// TIA Portal project "Parsing_migrated" (V16)

(* hardware
DEVICE "S71500/ET200MP station_1"  S7-1500 station
   slot 0: "Rail_0"  Rack  6ES7 590-1***0-0AA0
   slot 1: "PLC_1"  CPU 1515TF-2 PN  6ES7 515-2UM01-0AB0  V2.8
      slot 3: "CPU display_1"  6ES7591-1BA00-0AA0
      slot 32768: "PROFINET interface_1"  X1
         slot 32769: "Port_1"  X1 P1
         slot 32770: "Port_2"  X1 P2
      slot 33024: "PROFINET interface_2"  X2
         slot 33025: "Port_1"  X2 P1
      slot 34817: "Virtual CP interface port_1"  Virtual CP interface port  Virtual CP interface port
DEVICE "HMI_1"  KTP700F Mobile
   slot 0: "HMI_1"  KTP700F Mobile  6AV2 125-2GB23-0AX0  16.0.0.0
   slot 1: "HMI_RT_1"  KTP700F Mobile  6AV2 125-2GB23-0AX0  16.0.0.0
   slot 5: "HMI_1.IE_CP_1"  PROFINET Interface  16.0.0.0
      slot 1: "PROFINET Interface_1"  PROFINET Interface
         slot 1: "Port_1"  Port
DEVICE "SINAMICS S_1"  AcxSinamics.Device.2x.S210
   slot 0: "Left"  S210 PN  6SL3210-5HB10-1xFx  V5.2
      slot 1: "PROFINET interface"  PROFINET
      slot 3: " Ethernet commissioning interface"  LAN
   slot 0: "Drive control"  S210 PN
      slot 200: "Motor_Module_2"  Drive control  6SL3210-5HB10-1xFx
      slot 300: "SMIXX_3"  Drive control  1FK2102-1AG0x-xDAx
      slot 400: "Encoder_4"  Drive control  1FK2102-1AG0x-xDAx
      slot 1000: "Motor_SMI_5"  Drive control  1FK2102-1AG0x-xDAx
DEVICE "SINAMICS S_2"  AcxSinamics.Device.2x.S210
   slot 0: "Right"  S210 PN  6SL3210-5HB10-1xFx  V5.2
      slot 1: "PROFINET interface"  PROFINET
      slot 3: " Ethernet commissioning interface"  LAN
   slot 0: "Drive control"  S210 PN
      slot 200: "Motor_Module_2"  Drive control  6SL3210-5HB10-1xFx
      slot 300: "SMIXX_3"  Drive control  1FK2102-1AG0x-xDAx
      slot 400: "Encoder_4"  Drive control  1FK2102-1AG0x-xDAx
      slot 1000: "Motor_SMI_5"  Drive control  1FK2102-1AG0x-xDAx
*)

// ===== PLC "PLC_1"  CPU 1515TF-2 PN =====

VAR_GLOBAL   // PLC tag table "Default tag table"
   "PositioningAxis_Left_Actor_Interface_AddressIn" AT %I276.0 : "PD_TEL105_IN";
   "PositioningAxis_Left_Actor_Interface_AddressOut" AT %Q276.0 : "PD_TEL105_OUT";
   "PositioningAxis_Right_Actor_Interface_AddressIn" AT %I256.0 : "PD_TEL105_IN";
   "PositioningAxis_Right_Actor_Interface_AddressOut" AT %Q256.0 : "PD_TEL105_OUT";
   "actuator" AT %Q0.0 : Bool;
END_VAR

VAR_GLOBAL CONSTANT   // PLC tag table "LKinCtrl_PLC_Tags"
   "LKINCTRL_MC_MOVELINEARABS" : Int := 1;   // cmdType for linear absolute command
   "LKINCTRL_MC_MOVELINEARREL" : Int := 2;   // cmdType for linear relative command
   "LKINCTRL_MC_MOVECIRCULARABS" : Int := 3;   // cmdType for circular absolute command
   "LKINCTRL_MC_MOVECIRCULARREL" : Int := 4;   // cmdType for circular relative command
   "LKINCTRL_NO_OF_PATHDATA_PREBUFFER_ELEMENTS" : Int := 5;   // number of PreBuffer elements
   "LKINCTRL_NO_OF_START_EXECUTE_CMDS" : Int := 5;   // number of cmds to be buffered in first cycle
   "LKINCTRL_NO_OF_SEQ_EXECUTE_CMDS" : Int := 1;   // number of cmds to be buffered after first cycle
   "LKINCTRL_PI" : LReal := 3.1415926535897932846264;   // constant value for pi
   "LKINCTRL_NO_OF_CMD_SETFLAGS" : Int := 3;   // number of Boolean flags per command
   "LKINCTRL_LENGTH_OF_CMDPOINT_NAME" : Int := 10;   // length of point name
   "LKINCTRL_FM_SET_BEFORE_AND_NO_RESET" : USInt := 1;   // set flag before cmd and no reset
   "LKINCTRL_FM_SET_BEFORE_AND_RESET_AFTER" : USInt := 2;   // set flag before cmd and reset after
   "LKINCTRL_FM_SET_BEFORE_AND_RESET_AFTER_ONE_CYCLE" : USInt := 3;   // set flag before cmd and reset after one cycle
   "LKINCTRL_FM_SET_BEFORE_AND_NO_RESET_AND_WAIT_FOR_ACKNOWLEDGE" : USInt := 5;   // set flag before cmd and wait for external reset
   "LKINCTRL_FM_SET_AFTER_AND_NO_RESET" : USInt := 11;   // set flag after cmd and no reset
   "LKINCTRL_FM_SET_AFTER_AND_RESET_AFTER_ONE_CYCLE" : USInt := 13;   // set flag after cmd and reset after one cycle
   "LKINCTRL_FM_SET_AFTER_AND_NO_RESET_AND_WAIT_FOR_ACKNOWLEDGE" : USInt := 15;   // set flag after cmd and wait for external reset
   "LKINCTRL_FM_SET_AT_REMAINING_DISTANCE" : USInt := 10;   // set flag at remaining distance
   "LKINCTRL_FM_DISTANCE_TOLERANCE" : LReal := 0.01;   // tolerance for flagmode 10
   "LKINCTRL_NO_OF_SETFLAGS_BUFFER_ELEMENTS" : Int := 15;   // set as double of LKINCTRL_NO_OF_PATHDATA_PREBUFFER_ELEMENTS
   "LKINCTRL_COMP_LEFT" : Int := 1;   // tool radius compensation to the left
   "LKINCTRL_COMP_RIGHT" : Int := 2;   // tool radius compensation to the right
   "LKINCTRL_OUTER_CORNER" : Int := 1;   // Outer corner (linear / linear intersection)
   "LKINCTRL_INNER_CORNER" : Int := 2;   // Inner corner (linear / linear intersection)
   "LKINCTRL_CONFIG_END_OFFSET_COMP" : Int := 40;   // cmdType for ending offset compensation
   "LKINCTRL_CONFIG_START_OFFSET_COMP_LEFT" : Int := 41;   // cmdType for starting offset compensation left
   "LKINCTRL_NO_OF_PATHDATA_ELEMENTS" : Int := 20;   // length of LKinCtrl_typePathData
   "LKINCTRL_CMD_WAIT_TIME" : Int := 100;   // cmdType for wait time command
   "LKINCTRL_CONFIG_START_OFFSET_COMP_RIGHT" : Int := 42;   // cmdType for starting offset compensation right
   "LKINCTRL_LENGTH_OF_OFFSET_NAME" : Int := 10;   // length of offset name
   "LKINCTRL_NO_OF_OFFSETS" : Int := 3;   // number of configurable offsets
   "LKINCTRL_PATHDATA_TYPE_REDUCED" : USInt := 1;   // constant for PathData type "reduced"
   "LKINCTRL_PATHDATA_TYPE_NORMAL" : USInt := 2;   // constant for PathData type "normal"
   "LKINCTRL_PATHDATA_TYPE_ADVANCED" : USInt := 3;   // constant for PathData type "advanced"
   "LKINCTRL_NO_OF_PATHDATA_ELEMENTS_ADVANCED" : Int := 20;   // length of LKinCtrl_typePathData_advanced
   "LKINCTRL_NO_OF_PATHDATA_ELEMENTS_REDUCED" : Int := 10;   // length of LKinCtrl_typePathData_reduced
   "LKINCTRL_NO_OF_VALID_BITS" : Int := 4;   // number of valid bits in PathDataElement_advanced
   "LKINCTRL_CIRCMODE_GCODE" : Int := 3;   // circMode used in GCode
   "LKINCTRL_CMD_FLAG_ONLY" : Int := 0;   // cmdType for flagOnly command (no motion)
   "LKINCTRL_FM_DEACTIVATED" : USInt := 0;   // flag deactiavted
   "LKINCTRL_NO_OF_CMD_VALUEFLAGS" : Int := 3;   // number of LREAL flags per command
   "LKINCTRL_NO_OF_LAST_SETFLAG" : Int := 5;   // number of set flags at MovePath FB
   "LKINCTRL_NO_OF_LAST_VALUEFLAG" : Int := 5;   // number of value flags at MovePath FB
   "LKINCTRL_LENGTH_OF_PATHDATA_NAME" : Int := 15;   // length of PathData name
   "LKINCTRL_MC_MOVEDIRECTABS" : Int := 5;   // cmdType for move direct absolute command
   "LKINCTRL_MC_MOVEDIRECTREL" : Int := 6;   // cmdType for move direct relative command
   "LKINCTRL_NO_OF_CONVEYOR" : Int := 3;   // number of configurable offsets
   "LKINCTRL_MC_TRACKCONVEYORBELT" : Int := 10;   // cmdType for track conveyor belt command
END_VAR

VAR_GLOBAL CONSTANT   // PLC tag table "MC_Constants"
   "BM_BUFFERED" : Int := 1;   // Buffer mode 1: Standstill between motions
   "BM_BLENDING_LOW" : Int := 2;   // Buffer mode 2: Blending with lower velocity
   "BM_BLENDING_HIGH" : Int := 5;   // Buffer mode 5: Blending with higher velocity
   "DA_DEFAULT" : Int := -1;   // Dynamic adaption -1: Use default
   "DA_DEACTIVATED" : Int := 0;   // Dynamic adaption 0: Deactivated
   "DA_WITH_VARIABLE_LIMITS" : Int := 1;   // Dynamic adaption 1: With segmentation of path
   "DA_WITH_CONSTANT_LIMITS" : Int := 2;   // Dynamic adaption 2: No segmentation of path
   "SM_ACTIVE_DYNAMICS" : Int := 0;   // Stop mode 0: Stop with active dynamics
   "SM_MAX_DYNAMICS" : Int := 1;   // Stop mode 1: Stop with maximum dynamics
   "PC_POSITIVE" : Int := 0;   // Path choice 0: Shorter positive circle segment
   "PC_LONG_RUN_POSITIVE" : Int := 2;   // Path choice 2: Longer positive circle segment
   "PC_LONG_RUN_NEGATIVE" : Int := 3;   // Path choice 3: Longer negative circle segment
   "CP_XZ" : Int := 0;   // Circle plane 0: Circle in X-Z plane
   "CP_YZ" : Int := 1;   // Circle plane 1: Circle in Y-Z plane
   "CP_XY" : Int := 2;   // Circle plane 2: Circle in X-Y plane
   "CM_BORDER" : Int := 0;   // Circle mode 0: "EndPoint" + "AuxPoint" parameter defines a point on circular path
   "CM_CENTER" : Int := 1;   // Circle mode 1: "Arc" + "AuxPoint" defines circle center
   "CM_RADIUS" : Int := 2;   // Circle mode 2: "Radius" + "EndPoint" parameters define the circle segment
   "IM_ACTIVE_DYNAMICS" : Int := 0;   // Interrupt mode 0: Interrupt with active dynamics
   "IM_MAX_DYNAMICS" : Int := 1;   // Interrupt mode 1: Interrupt with maximum dynamics
   "DIRA_POSITIVE" : Int := 1;   // Orientation direction 1: Positive direction
   "DIRA_NEGATIVE" : Int := 2;   // Orientation direction 2: Negative direction
   "DIRA_SHORTEST" : Int := 3;   // Orientation direction 3: Shortest direction
   "CS_WCS" : Int := 0;   // Coordinate system 0: World coordinate system (WCS)
   "CS_OCS1" : Int := 1;   // Coordinate system 1: Object coordinate system 1 (OCS[1])
   "CS_OCS2" : Int := 2;   // Coordinate system 2: Object coordinate system 2 (OCS[2])
   "CS_OCS3" : Int := 3;   // Coordinate system 3: Object coordinate system 3 (OCS[3])
   "PC_NEGATIVE" : Int := 1;   // Path choice 1: Shorter negative circle segment
   "CS_MCS" : Int := 100;   // Coordinate system 100: Machine coordinate system (axis values)
   "LC_DEFAULT" : DWord := 16#FFFFFFFF;   // LinkConstellation: Default to keep link constellation of kinematics
   "PM_ABS_ABS" : DInt := 1;   // PositionMode 1: Interpretation of cartesian orientation as absolute (only effective for absolute MoveDirect commands)
   "PM_ABS_REL" : DInt := 2;   // PositionMode 2: Interpretation of cartesian orientation as relative (only effective for absolute MoveDirect commands)
END_VAR

VAR_GLOBAL CONSTANT   // PLC tag table "LKinLang_Configuration"
   "LKINLANG_FIRST_INDEX_LINE_BUFFER" : Int := 1;   // First index of the line buffer
   "LKINLANG_LAST_INDEX_LINE_BUFFER" : Int := 20;   // Last index of the line buffer
   "LKINLANG_LENGTH_OF_ASCII_LINE_STRING" : UDInt := 128;   // Maximum number of ASCII characters in one line (without CR/LF)
   "LKINLANG_LENGTH_OF_TOKEN_STRING" : Int := 20;   // Maximum string length of one token
   "LKINLANG_MAX_NUMBER_OF_TOKEN_PER_LINE" : Int := 50;   // Maximum number of token per line
   "LKINLANG_MAX_NUMBER_OF_PARAMETERS_PER_LINE" : Int := 25;   // Maximum number of parameters in one line
   "LKINLANG_MAX_NUMBER_OF_PARAMETERS" : Int := 125;   // Maximum number of configured language parameters (G1,G2,...)
   "LKINLANG_NUMBER_OF_SEPARATORS" : Int := 15;   // Maximum number of separators
   "LKINLANG_NUMBER_OF_MERGERS" : Int := 10;   // Maximum number of mergers
   "LKINLANG_NUMBER_OF_FOLLOW_VALUES" : Int := 4;   // Maximum number of follow values for one command
   "LKINLANG_NUMBER_OF_CONDITIONS" : Int := 50;   // Maximum number of conditions for one command
   "LKINLANG_NUMBER_OF_REPLACEMENTS" : Int := 10;   // Maximum number of replacements
   "LKINLANG_NUMBER_OF_LABELS" : Int := 20;   // Maximum number of labels
   "LKINLANG_NUMBER_OF_STACK_ELEMENTS" : Int := 20;   // Maximum number of stack elements
   "LKINLANG_NUMBER_OF_HIERARCHICLEVEL" : Int := 60;   // Maximum number of hierarchic level changes
   "LKINLANG_NUMBER_OF_SUBPROGRAMS" : Int := 10;   // Maximum number of subprograms
   "LKINLANG_NUMBER_OF_VAR_REFS" : Int := 20;   // Maximum number of variable references
   "LKINLANG_NUMBER_OF_INTERFACE_BOOL" : Int := 5;   // Maximum number of boolean interface variables
   "LKINLANG_NUMBER_OF_INTERFACE_DINT" : Int := 10;   // Maximum number of DInt interface variables
   "LKINLANG_NUMBER_OF_INTERFACE_LREAL" : Int := 20;   // Maximum number of LReal interface variables
   "LKINLANG_NUMBER_OF_LOCAL_BOOL" : Int := 10;   // Maximum number of boolean local variables
   "LKINLANG_NUMBER_OF_LOCAL_DINT" : Int := 10;   // Maximum number of DInt local variables
   "LKINLANG_NUMBER_OF_LOCAL_LREAL" : Int := 10;   // Maximum number of LReal local variables
   "LKINLANG_LANGPACK_GCODE" : Int := 1;   // Select GCode language package
   "LKINLANG_LANGPACK_USER" : Int := 2;   // Select user defined language package
END_VAR

VAR_GLOBAL CONSTANT   // PLC tag table "LKinLang_Constants"
   "LKINLANG_PRIO_UNRELEVANT" : Int := 0;   // Lowest parameter priority
   "LKINLANG_PRIO_DEFAULT" : Int := 1;   // Normal parameter priority
   "LKINLANG_PRIO_DEFINED" : Int := 2;   // High parameter priority
   "LKINLANG_PRIO_CONSTANT" : Int := 3;   // Highest parameter priority
   "LKINLANG_MOTION_CMD" : DWord := 2#0000_0001;   // Parameter property: Motion command
   "LKINLANG_ABSOLUTE_POSITION" : DWord := 2#0010_0000;   // Parameter property: Switch to absolute positioning
   "LKINLANG_RELATIVE_POSITION" : DWord := 2#0100_0000;   // Parameter property: Switch to relative positioning
   "LKINLANG_CMD_MODAL" : DWord := 2#0000_0010;   // Parameter property: Modal until change of motion command
   "LKINLANG_PRG_MODAL" : DWord := 2#0000_0100;   // Parameter property: Modal for complete program
   "LKINLANG_CHECK_LIMITS" : DWord := 2#0000_1000;   // Parameter property: Check limits for parameter
   "LKINLANG_EQUATION" : DWord := 2#0001_0000;   // Parameter property: Math expressions allowed
   "LKINLANG_CONDITION_IN_LINE" : DInt := 1;   // Condition check: Condition must be set in same line
   "LKINLANG_CONDITION_IN_COMMAND" : DInt := 2;   // Condition check: Condition must be set in same motion command
   "LKINLANG_CONDITION_IN_PROGRAM" : DInt := 3;   // Condition check: Condition must be set in program before
   "LKINLANG_FILE_STATE_RUNNING" : DInt := 200;   // File status: Program in execution
   "LKINLANG_FILE_STATE_STOPPED" : DInt := 90;   // File status: Program stopped
   "LKINLANG_FILE_STATE_EDITING" : DInt := 20;   // File status: Program is edited
   "LKINLANG_FILE_STATE_LOADING" : DInt := 10;   // File status: Program is being loaded from MMC
   "LKINLANG_FILE_STATE_RUNNING_LOADING" : DInt := 300;   // File status: Program is executed and loaded simultaneously
   "LKINLANG_FILE_STATE_SAVING" : DInt := 30;   // File status: Program is being saved
   "LKINLANG_FILE_STATE_IDLE" : DInt := 100;   // File status: Program is ready
   "LKINLANG_FILE_STATE_SAVE_REQUESTED" : DInt := 40;   // File status: Program saving is requested
   "LKINLANG_VAR_TYPE_LOCAL_BOOL" : Int := 1;   // Type constant for local boolean variables
   "LKINLANG_VAR_TYPE_LOCAL_DINT" : Int := 2;   // Type constant for local integer variables
   "LKINLANG_VAR_TYPE_LOCAL_LREAL" : Int := 3;   // Type constant for local real variables
   "LKINLANG_VAR_TYPE_INTERFACE_BOOL" : Int := 101;   // Type constant for boolean interface variables
   "LKINLANG_VAR_TYPE_INTERFACE_DINT" : Int := 102;   // Type constant for integer interface variables
   "LKINLANG_VAR_TYPE_INTERFACE_LREAL" : Int := 103;   // Type constant for real interface variables
   "LKINLANG_SYNTAX_CHECK_OFF" : USInt := 0;   // Constant for syntax check: No check before writing commands
   "LKINLANG_SYNTAX_CHECK_ONLY" : USInt := 1;   // Constant for syntax check: Only check; no writing of commands
   "LKINLANG_SYNTAX_CHECK_AND_EXECUTE" : USInt := 2;   // Constant for syntax check: Check before and write commands after check
   "LKINLANG_ENTRY_TYPE_IF" : Int := 10;   // Stack entry type IF
   "LKINLANG_ENTRY_TYPE_ELSE" : Int := 11;   // Stack entry type ELSE
   "LKINLANG_ENTRY_TYPE_ENDIF" : Int := 12;   // Stack entry type ENDIF
   "LKINLANG_ENTRY_TYPE_WHILE" : Int := 20;   // Stack entry type WHILE
   "LKINLANG_ENTRY_TYPE_ENDWHILE" : Int := 22;   // Stack entry type ENDWHILE
   "LKINLANG_ENTRY_TYPE_FOR" : Int := 30;   // Stack entry type FOR
   "LKINLANG_ENTRY_TYPE_ENDFOR" : Int := 32;   // Stack entry type ENDFOR
   "LKINLANG_ENTRY_TYPE_SUB" : Int := 40;   // Stack entry type SUB
END_VAR

// folder: LKinCtrl_Types

TYPE "LKinCtrl_typeFrame"
   STRUCT
      x : LReal;   // Translation in x
      y : LReal;   // Translation in y
      z : LReal;   // Translation in z
      "a" : LReal;   // Rotation around z axis
      "b" : LReal;   // Rotation around y axis
      c : LReal;   // Roataion around x axis
   END_STRUCT;
END_TYPE

TYPE "LKinCtrl_typePathDataElement_advanced"
VERSION : 0.1
   STRUCT
      cmdType : Int := -1;   // 1: MoveLinAbs; 2: MoveLinRel; 3: MoveCircAbs; 4: MoveCircRel; 5: MoveDirectAbs; 6: MoveDirectRel; 10: TrackConveyorBelt; 100: WaitTime; 40/41/42: ContourOffset; 0: FlagOnlyCmd; -1: End of List
      cmdActivated : Bool := TRUE;   // (de)activation of command
      cmdName : String["LKINCTRL_LENGTH_OF_CMDPOINT_NAME"];   // name of command
      cmdCoordinates : "LKinCtrl_typePointCoordinates";   // target coordinate definition
      cmdParameters : "LKinCtrl_typePointParameter";   // additional command parameters
      setFlags : Array[1.."LKINCTRL_NO_OF_CMD_SETFLAGS"] of "LKinCtrl_typeSetFlagElement_Bool";   // flags to control actuators
      valueFlags : Array[1.."LKINCTRL_NO_OF_CMD_VALUEFLAGS"] of "LKinCtrl_typeSetFlagElement_LReal";   // value flags to control actuators
      parameterValid : Array[1..4] of Bool;   // valid bit for cartesian position parameters
   END_STRUCT;
   // parameterValid[1] := True;   // X
   // parameterValid[2] := True;   // Y
   // parameterValid[3] := True;   // Z
   // parameterValid[4] := True;   // A
   // // cmdParameters.transitionParameters : blending parameters
   // // cmdParameters.pathDynamics : dynamic settings
END_TYPE

TYPE "LKinCtrl_typeCmdLoggerElement"
VERSION : 0.1
   STRUCT
      cmdType : Int := -1;   // 1: MoveLinAbs; 2: MoveLinRel; 3: MoveCircAbs; 4: MoveCircRel; 5: MoveDirectAbs; 6: MoveDirectRel; 10: TrackConveyorBelt; 100: WaitTime; 40/41/42: ContourOffset; 0: FlagOnlyCmd; -1: End of List
      pathDataName : String["LKINCTRL_LENGTH_OF_PATHDATA_NAME"];   // name of PathData
      pathDataIdentifier : Int;   // identifier of PathData containing command
      cmdID : DInt;   // to be set to PathDataOperate[list position] by PreBuffer for identification in ExecuteBuffer
      cmdName : String[4];   // command name
      coordinateX : LReal;   // X (linear) / endPoint[1] (circular)
      coordinateY : LReal;   // Y (linear) / endPoint[2] (circular)
      coordinateZ : LReal;   // Z (linear) / endPoint[3] (circular)
      coordinateA : LReal;   // A (linear) / endPoint[4] (circular)
      coordSystem : DInt := 0;   // 0: WCS; 1: OCS[1]; 2: OCS[2]; 3: OCS[3]
      bufferMode : DInt := 1;   // 1: standstill between commands, 2: blending with lower speed; 5: blending with higher speed
      transitionParameter : LReal;   // blending distance - >0.0: configured value used; <0.0: maximum possible blending distance used
      dynVelocity : LReal;   // >0.0: configured value used; <0.0: default TO setting used
      dynAcceleration : LReal;   // >0.0: configured value used; <0.0: default TO setting used
      dynDeceleration : LReal;   // >0.0: configured value used; <0.0: default TO setting used
      dynJerk : LReal;   // >0.0: configured value used; <0.0: default TO setting used
      dynamicAdpation : DInt;   // <0.0: default TO setting used; 0: no dynamic adaption; 1: with variable limits; 2: with constant limits
      linkConstellation : DWord;   // linkConstellation (effective for MoveDirect commands only)
      positionMode : DInt;   // 1: absolute cartesian position and absolute orientation; 2: absolute cartesian position and relative orientation (effective for MoveDirect commands only)
      circMode : DInt;   // 0: auxPoint defines point on circle line; 1: auxPoint defines circle center; 2: radius and endPoint define circle segment
      auxPoint_1 : LReal;   // auxiliary point for circle definition
      auxPoint_2 : LReal;   // auxiliary point for circle definition
      auxPoint_3 : LReal;   // auxiliary point for circle definition
      pathChoice : DInt;   // circMode(0): not relevant; circMode(1): 0: pos direction; 1: neg direction; circMode(2): 0: short pos segment; 1: short neg segment; 2: long pos segment; 3: long neg segment
      circlePlane : DInt;   // circMode(0): not relevant; circMode(1+2): 0: XZ; 1: YZ; 2: XY
      radius : LReal;   // only in combination with circMode(2): radius
      arc : LReal;   // only in combination with circMode(1): arc
   END_STRUCT;
END_TYPE

TYPE "LKinCtrl_typeSetFlagElement_LReal"
VERSION : 0.1
   STRUCT
      flag : Int := -1;   // index of flag to be set
      value : LReal := 0.0;   // value for flagValue
      flagMode : USInt := 1;   // (see LKinCtrl_PLC_Tags) 0: deactivated; 1: SET_BEFORE_AND_NO_RESET; 2: SET_BEFORE_AND_RESET_AFTER; 3: SET_BEFORE_AND_RESET_AFTER_ONE_CYCLE; 5: SET_BEFORE_AND_NO_RESET_AND_WAIT_FOR_ACKNOWLEDGE; 10: LKINCTRL_FM_SET_AT_REMAINING_DISTANCE; 11: LKINCTRL_FM_SET_AFTER_AND_NO_RESET; 13: LKINCTRL_FM_SET_AFTER_AND_RESET_AFTER_ONE_CYCLE; 15: LKINCTRL_FM_SET_AFTER_AND_NO_RESET_AND_WAIT_FOR_ACKNOWLEDGE
      remainingDistance : LReal := -1.0;   // >0.0: remainingDistance
   END_STRUCT;
END_TYPE

TYPE "LKinCtrl_typeSetFlagElement_Bool"
VERSION : 0.1
   STRUCT
      flag : Int := -1;   // flag to be set
      flagMode : USInt := 1;   // (see LKinCtrl_PLC_Tags) 0: deactivated; 1: SET_BEFORE_AND_NO_RESET; 2: SET_BEFORE_AND_RESET_AFTER; 3: SET_BEFORE_AND_RESET_AFTER_ONE_CYCLE; 5: SET_BEFORE_AND_NO_RESET_AND_WAIT_FOR_ACKNOWLEDGE; 10: LKINCTRL_FM_SET_AT_REMAINING_DISTANCE; 11: LKINCTRL_FM_SET_AFTER_AND_NO_RESET; 13: LKINCTRL_FM_SET_AFTER_AND_RESET_AFTER_ONE_CYCLE; 15: LKINCTRL_FM_SET_AFTER_AND_NO_RESET_AND_WAIT_FOR_ACKNOWLEDGE
      remainingDistance : LReal := -1.0;   // >0.0: remainingDistance
   END_STRUCT;
END_TYPE

TYPE "LKinCtrl_typePointCoordinates"
VERSION : 0.1
   STRUCT
      cartesianPosition : "LKinCtrl_typeCartesianPosition";   // cartesian position
      coordSystem : DInt := 0;   // 0: WCS; 1: OCS[1]; 2: OCS[2]; 3: OCS[3] / 0: WCS; 1: OCS[1]; 2: OCS[2]; 3: OCS[3]; 100: MCS
   END_STRUCT;
END_TYPE

TYPE "LKinCtrl_typePointCoordinates_PreBuf"
VERSION : 0.1
   STRUCT
      absolutePosition : Array[1..4] of LReal;   // absolute cartesian position
      coordSystem : DInt := 0;   // 0: WCS; 1: OCS[1]; 2: OCS[2]; 3: OCS[3]
   END_STRUCT;
   // // absolutePosition[1] : X
   // // absolutePosition[2] : Y
   // // absolutePosition[3] : Z
   // // absolutePosition[4] : A
END_TYPE

TYPE "LKinCtrl_typePathDynamics"
VERSION : 0.1
   STRUCT
      velocity : LReal := -1.0;   // >0.0: configured value used; <0.0: default TO setting used; for cmdType = 100 ==> waitTime in ms
      acceleration : LReal := -1.0;   // >0.0: configured value used; <0.0: default TO setting used
      deceleration : LReal := -1.0;   // >0.0: configured value used; <0.0: default TO setting used
      jerk : LReal := -1.0;   // >0.0: configured value used; <0.0: default TO setting used
   END_STRUCT;
END_TYPE

TYPE "LKinCtrl_typePathDataElement_PreBuf"
VERSION : 0.1
   STRUCT
      cmdType : Int := -1;   // 1: MoveLinAbs; 2: MoveLinRel; 3: MoveCircAbs; 4: MoveCircRel; 5: MoveDirectAbs; 6: MoveDirectRel; 10: TrackConveyorBelt; 100: WaitTime; 40/41/42: ContourOffset; 0: FlagOnlyCmd; -1: End of List
      cmdID : DInt;   // to be set to PathDataOperate[list position] by PreBuffer for identification in ExecuteBuffer
      cmdName : String["LKINCTRL_LENGTH_OF_CMDPOINT_NAME"];   // command name
      cmdCoordinates : "LKinCtrl_typePointCoordinates_PreBuf";   // command coordinates
      cmdParameters : "LKinCtrl_typePointParameter";   // command parameters
      pathDataName : String["LKINCTRL_LENGTH_OF_PATHDATA_NAME"];   // name of PathData
      pathDataIdentifier : USInt;   // identifier of PathData
      isIntermediateCmd : Bool;   // TRUE: command is intermediate command
      setFlags : Array[1.."LKINCTRL_NO_OF_CMD_SETFLAGS"] of "LKinCtrl_typeSetFlagElement_Bool";   // flags to control actuators
      valueFlags : Array[1.."LKINCTRL_NO_OF_CMD_VALUEFLAGS"] of "LKinCtrl_typeSetFlagElement_LReal";   // value flags to control actuators
      parameterValid : Array[1..4] of Bool;   // valid bit for cartesian position parameters
   END_STRUCT;
   // parameterValid[1] := True;   // X
   // parameterValid[2] := True;   // Y
   // parameterValid[3] := True;   // Z
   // parameterValid[4] := True;   // A
END_TYPE

TYPE "LKinCtrl_typePathDescriptionElement"
   STRUCT
      pointName : String["LKINCTRL_LENGTH_OF_CMDPOINT_NAME"];   // name of point
      targetPosition : "LKinCtrl_typeCartesianPosition";   // target position
      coordSystem : DInt;   // 0: WCS; 1: OCS[1]; 2: OCS[2]; 3: OCS[3]
      blendingDistance : LReal;   // blending radius
      flags : Array[1.."LKINCTRL_NO_OF_CMD_SETFLAGS"] of "LKinCtrl_typeSetFlagElement_Bool";   // flags to control actuators
      valueFlags : Array[1.."LKINCTRL_NO_OF_CMD_VALUEFLAGS"] of "LKinCtrl_typeSetFlagElement_LReal";   // value flags to control actuators
   END_STRUCT;
END_TYPE

TYPE "LKinCtrl_typePointParameter"
VERSION : 0.1
   STRUCT
      pathDynamics : "LKinCtrl_typePathDynamics";   // dynamics settings for single command
      orientationDirection : DInt := 3;   // 1: positive direction; 2: negative direction; 3: shortest distance
      bufferMode : DInt := 1;   // 1: standstill between commands, 2: blending with lower speed; 5: blending with higher speed
      transitionParameters : Array[1..5] of LReal;   // blending distance parameters
      dynamicAdaption : DInt := -1;   // <0.0: default TO setting used; 0: no dynamic adaption; 1: with variable limits; 2: with constant limits
      moveDirectParameters : "LKinCtrl_typeMoveDirectParameter";   // parameters for MoveDirect command definition
      offsetParameters : "LKinCtrl_typeToolParameters";   // parameters for offset selection and configuration
      conveyorParameters : "LKinCtrl_typeConveyorParameter";   // parameters for conveyor selection and configuration
      circleParameters : "LKinCtrl_typeCircleParameters";   // parameters for circle command definition
   END_STRUCT;
   // transitionParameters[1] := -1.0;   // blending distance - >0.0: configured value used; <0.0: maximum possible blending distance used
   // // transitionParameters[2] : reserved, do not set
   // // transitionParameters[3] : reserved, do not set
   // // transitionParameters[4] : reserved, do not set
   // // transitionParameters[5] : reserved, do not set
END_TYPE

TYPE "LKinCtrl_typePathData_advanced"
VERSION : 0.1
   STRUCT
      pathDataName : String["LKINCTRL_LENGTH_OF_PATHDATA_NAME"];   // name of PathData
      pointers : "LKinCtrl_typeAdvPointers";   // pointers to add / retrieve cmds in PathData
      commands : Array[1.."LKINCTRL_NO_OF_PATHDATA_ELEMENTS_ADVANCED"] of "LKinCtrl_typePathDataElement_advanced";   // command list
   END_STRUCT;
END_TYPE

TYPE "LKinCtrl_typePathDataElement"
VERSION : 0.1
   STRUCT
      cmdType : Int := -1;   // 1: MoveLinAbs; 2: MoveLinRel; 3: MoveCircAbs; 4: MoveCircRel; 5: MoveDirectAbs; 6: MoveDirectRel; 10: TrackConveyorBelt; 100: WaitTime; 40/41/42: ContourOffset; 0: FlagOnlyCmd; -1: End of List
      cmdActivated : Bool := TRUE;   // (de)activation of command
      cmdName : String["LKINCTRL_LENGTH_OF_CMDPOINT_NAME"];   // name of command
      cmdCoordinates : "LKinCtrl_typePointCoordinates";   // target coordinate definition
      cmdParameters : "LKinCtrl_typePointParameter";   // additional command parameters
      setFlags : Array[1.."LKINCTRL_NO_OF_CMD_SETFLAGS"] of "LKinCtrl_typeSetFlagElement_Bool";   // flags to control actuators
      valueFlags : Array[1.."LKINCTRL_NO_OF_CMD_VALUEFLAGS"] of "LKinCtrl_typeSetFlagElement_LReal";   // value flags to control actuators
   END_STRUCT;
   // // cmdParameters.transitionParameters : blending parameters
   // // cmdParameters.pathDynamics : dynamic settings
END_TYPE

TYPE "LKinCtrl_typePathDescription"
   STRUCT
      pathDescriptionName : String[10];   // name of PathDescription
      points : Array[1.."LKINCTRL_NO_OF_PATHDATA_ELEMENTS"] of "LKinCtrl_typePathDescriptionElement";   // target points
   END_STRUCT;
END_TYPE

TYPE "LKinCtrl_typeAdvPointers"
VERSION : 0.1
   STRUCT
      addPointer : DInt := 0;   // pointer to add new comds to PathData after cmd has been executed by MovePath
      retrievePointer : DInt := 0;   // pointer to show which cmd is the next to be retrieved by MovePath
      addPointerRestarted : Bool;   // addPointer restarted after overflow
      ignoreAddPointer : Bool := true;   // addPointer not taken into account for buffering, unless set by previous data source
      bufferLocked : Bool;   // buffer locked to wait for previous data source - read data locked
      preprocessingStop : Bool;   // parser reached a preprocessing stop
   END_STRUCT;
END_TYPE

TYPE "LKinCtrl_typePointParameter_reduced"
VERSION : 0.1
   STRUCT
      pathDynamics : "LKinCtrl_typePathDynamics";   // dynamics settings for single command
      orientationDirection : DInt := 3;   // 1: positive direction; 2: negative direction; 3: shortest distance
      bufferMode : DInt := 1;   // 1: standstill between commands, 2: blending with lower speed; 5: blending with higher speed
      transitionParameters : Array[1..5] of LReal;   // blending distance parameters
      dynamicAdaption : DInt := -1;   // <0.0: default TO setting used; 0: no dynamic adaption; 1: with variable limits; 2: with constant limits
   END_STRUCT;
   // transitionParameters[1] := -1.0;   // blending distance - >0.0: configured value used; <0.0: maximum possible blending distance used
   // // transitionParameters[2] : reserved, do not set
   // // transitionParameters[3] : reserved, do not set
   // // transitionParameters[4] : reserved, do not set
   // // transitionParameters[5] : reserved, do not set
END_TYPE

TYPE "LKinCtrl_typePathData_reduced"
VERSION : 0.1
   STRUCT
      pathDataName : String["LKINCTRL_LENGTH_OF_PATHDATA_NAME"];   // name of PathData
      commands : Array[1.."LKINCTRL_NO_OF_PATHDATA_ELEMENTS_REDUCED"] of "LKinCtrl_typePathDataElement_reduced";   // command list
   END_STRUCT;
END_TYPE

TYPE "LKinCtrl_typePathData"
VERSION : 0.1
   STRUCT
      pathDataName : String["LKINCTRL_LENGTH_OF_PATHDATA_NAME"];   // name of PathData
      commands : Array[1.."LKINCTRL_NO_OF_PATHDATA_ELEMENTS"] of "LKinCtrl_typePathDataElement";   // command list
   END_STRUCT;
END_TYPE

TYPE "LKinCtrl_typePathData_PreBuf"
VERSION : 0.1
   STRUCT
      pathDataName : String["LKINCTRL_LENGTH_OF_PATHDATA_NAME"];   // name of PathData
      commands : Array[1.."LKINCTRL_NO_OF_PATHDATA_PREBUFFER_ELEMENTS"] of "LKinCtrl_typePathDataElement_PreBuf";   // command list
      addPointer : Int;   // pointer marking slot for adding of next command in PathDataPreBuffered
      retrievePointer : Int;   // pointer marking command entry to be read in PathDataPreBuffered
      addPointerRestarted : Bool;   // addPointer restarted after overflow
   END_STRUCT;
END_TYPE

TYPE "LKinCtrl_typePathDataElement_reduced"
VERSION : 0.1
   STRUCT
      cmdType : Int := -1;   // 1: MoveLinAbs; 2: MoveLinRel; 100: WaitTime; 0: FlagOnlyCmd; -1: End of List
      cmdActivated : Bool := TRUE;   // (de)activation of command
      cmdName : String["LKINCTRL_LENGTH_OF_CMDPOINT_NAME"];   // name of command
      cmdCoordinates : "LKinCtrl_typePointCoordinates";   // target coordinate definition
      cmdParameters : "LKinCtrl_typePointParameter_reduced";   // additional command parameters
      setFlags : Array[1.."LKINCTRL_NO_OF_CMD_SETFLAGS"] of "LKinCtrl_typeSetFlagElement_Bool";   // flags to control actuators
      valueFlags : Array[1.."LKINCTRL_NO_OF_CMD_VALUEFLAGS"] of "LKinCtrl_typeSetFlagElement_LReal";   // value flags to control actuators
   END_STRUCT;
END_TYPE

TYPE "LKinCtrl_typeDiagnosticsPathSelect"
TITLE = typeDiagnosticsFBTemplate
VERSION : 0.1
   STRUCT
      status : Word;   // Status of the FC or error identification when error occurred
      entryID : Int;   // identifier for false entry
   END_STRUCT;
END_TYPE

TYPE "LKinCtrl_typeExecuteKinMotionCmdDiagnostics"
VERSION : 0.1
   STRUCT
      status : Word;   // status of the FB
      faultPathDataName : String["LKINCTRL_LENGTH_OF_PATHDATA_NAME"];   // number of PathData with occurring error in PathData set
      faultSetNumber : DInt;   // number of PathData set with occurring error
      faultFBNumber : DInt;   // number of motionCommand FB with occurring error
      motionFBstatus : DWord;   // status of motion FB (internal) an error occurred in
      stateMachine : Int;   // stateMachine status
      kinematicsStatusWord : DWord;   // statusWord TO kinematics
      kinematicsErrorWord : DWord;   // errorWord TO kinematics
   END_STRUCT;
END_TYPE

TYPE "LKinCtrl_typeCircleParameters"
VERSION : 0.1
   STRUCT
      circMode : DInt := 0;   // 0: auxPoint defines point on circle line; 1: auxPoint defines circle center; 2: radius and endPoint define circle segment; 3: GCode notation (end & aux point)
      auxPoint : Array[1..3] of LReal;   // auxiliary point for circle definition
      pathChoice : DInt := 0;   // circMode(0): not relevant; circMode(1): 0: pos direction; 1: neg direction; circMode(2): 0: short pos segment; 1: short neg segment; 2: long pos segment; 3: long neg segment
      circlePlane : DInt;   // circMode(0): not relevant; circMode(1+2): 0: XZ; 1: YZ; 2: XY
      radius : LReal;   // only in combination with circMode(2): radius
      arc : LReal;   // only in combination with circMode(1): arc
   END_STRUCT;
   // // auxPoint[1] : X
   // // auxPoint[2] : Y
   // // auxPoint[3] : Z
END_TYPE

TYPE "LKinCtrl_typeMovePathDiagnostics"
VERSION : 0.1
   STRUCT
      errorID : Word;   // errorID of the FB
      pathDataName : String["LKINCTRL_LENGTH_OF_PATHDATA_NAME"];   // name of PathData an error occurred in
      cmdNumber : DInt;   // command number (in PathData) an error occurred in
      stateMovePath : DInt;   // state machine status FB
      statusSubFunction : Word;   // status of LKinCtrl_MC_ExecuteKinMotionCmd
      motionFBNumber : DInt;   // motion FB number (internal) an error occurred in
      motionFBStatus : DWord;   // status of motion FB (internal) an error occurred in
      kinematicsStatusWord : DWord;   // statusWord TO kinematics
      kinematicsErrorWord : DWord;   // errorWord TO kinematics
   END_STRUCT;
END_TYPE

TYPE "LKinCtrl_typeJogFrameDiagnostics"
VERSION : 0.1
// support: tech.team.motioncontrol@siemens.com
   STRUCT
      timeStamp : Date_And_Time;   // Time stamp at which the error occurred
      status : Word;   // Status of FB when error occurred
      stateNumber : DInt;   // State in the state machine of the FB when the error occurred
   END_STRUCT;
END_TYPE

TYPE "LKinCtrl_typeCartesianPosition"
VERSION : 0.1
   STRUCT
      x : LReal;   // X
      y : LReal;   // Y
      z : LReal;   // Z
      "a" : LReal;   // A
   END_STRUCT;
END_TYPE

TYPE "LKinCtrl_typeDynamics"
VERSION : 0.1
   STRUCT
      path : "LKinCtrl_typePathDynamics";   // Specification of the path dynamics
      orientation : "LKinCtrl_typePathDynamics";   // Specification of the orientation dynamics
      dynamicAdaption : DInt := 1;   // 0=no dynamic adaption, 1=dynamic adaptation with segmentation of the path, 2=dynamic adaptation without segmentation of the path
   END_STRUCT;
END_TYPE

TYPE "LKinCtrl_typeAuxFCDiagnostics"
TITLE = typeDiagnosticsFBTemplate
   STRUCT
      status : Word;   // Status of the FB or error identification when error occurred
      subfunctionStatus : Word;   // Status or return value of called FBs, FCs and system blocks
      axisNumber : Int;   // number of the corresponding axis the error occured in or a function effecting it
      errorDetail : UDInt;   // error detail of corresponding technology object the error occured in
      stateNumber : DInt;   // State in the state machine of the FB when the error occurred
   END_STRUCT;
END_TYPE

TYPE "LKinCtrl_typeMoveDirectParameter"
VERSION : 0.1
   STRUCT
      linkConstellation : DWord := 16#FFFFFFFF;   // linkConstellation (effective for MoveDirect commands only)
      positionMode : DInt := 1;   // 1: absolute cartesian position and absolute orientation; 2: absolute cartesian position and relative orientation (effective for MoveDirect commands only)
   END_STRUCT;
END_TYPE

TYPE "LKinCtrl_typeConfiguration"
   STRUCT
      offsetParameter : Array[1.."LKINCTRL_NO_OF_OFFSETS"] of "LKinCtrl_typeContourOffsetParameter";   // offset parameter settings
      conveyorParameter : Array[1.."LKINCTRL_NO_OF_CONVEYOR"] of "LKinCtrl_typeConveyorConfiguration";   // conveyor parameter settings
      stopMode : DInt;   // MC_GroupStop dynamics; 0: stop with dynamics of active motion job; 1: stop with maximum kinematics dynamics (dynamics adaption still effective); 10: stop with dynamics of active motion job and desync conveyor; 11: stop with maximum kinematics dynamics and desync conveyor
   END_STRUCT;
END_TYPE

TYPE "LKinCtrl_typeContourOffsetParameter"
   STRUCT
      "name" : String["LKINCTRL_LENGTH_OF_OFFSET_NAME"];   // offset name
      radius : LReal;   // offset radius
      length : LReal;   // offset length
   END_STRUCT;
END_TYPE

TYPE "LKinCtrl_typeToolParameters"
   STRUCT
      offsetParaNo : Int;   // selection of offset parameter set from configuration structure
      mainPathPlane : Int;   // main path plane for compensation
   END_STRUCT;
END_TYPE

TYPE "LKinCtrl_typeConveyorParameter"
   STRUCT
      conveyorParaNo : DInt := 1;   // selection of conveyor parameter set from configuration structure
   END_STRUCT;
END_TYPE

TYPE "LKinCtrl_typeConveyorConfiguration"
   STRUCT
      conveyorBeltAxis : DB_ANY;   // Conveyor belt axis DB
      conveyorBeltOrigin : TO_Struct_Kinematics_Frame;   // Frane to origin of conveyor belt
      initialObjectPosition : TO_Struct_Kinematics_Frame;   // Initial object position on conveyor (only x allowed)
   END_STRUCT;
END_TYPE

// folder: LKinCtrl_Types/LKinCtrl_ContOffset_Types

TYPE "LKinCtrl_typeCOff3DPoint"
VERSION : 0.1
   STRUCT
      x : LReal;   // X
      y : LReal;   // Y
      z : LReal;   // Z
   END_STRUCT;
END_TYPE

TYPE "LKinCtrl_typeCOffReturn"
   STRUCT
      returnValue : Word;   // Return value
      region : Int;   // Region type - see LKinCtrl_OffsetContour
      subBlockNumber : DInt;   // Sub function block number
      internalNumber : DInt;   // Internal number indicates the source code position
   END_STRUCT;
END_TYPE

TYPE "LKinCtrl_typeCOffPathDataIn"
   STRUCT
      currentPos : "LKinCtrl_typeCOffInCurrentPos";   // Source data - current position
      nextCommand : "LKinCtrl_typePathDataElement";   // Source data - next command
      nextButOneCommand : "LKinCtrl_typePathDataElement";   // Source data - next but one command
   END_STRUCT;
END_TYPE

TYPE "LKinCtrl_typeCOffOutNextButOneCmd"
   STRUCT
      transitionParameter : Array[1..5] of LReal;   // blending parameters
   END_STRUCT;
END_TYPE

TYPE "LKinCtrl_typeCOffCmdInInternal"
   STRUCT
      cmdType : Int := -1;   // 1: MoveLinAbs; 2: MoveLinRel; 3: MoveCircAbs; 4: MoveCircRel; 5: MoveDirectAbs; 6: MoveDirectRel; 10: TrackConveyorBelt; 100: WaitTime; 40/41/42: ContourOffset; 0: FlagOnlyCmd; -1: End of List
      endPoint : "LKinCtrl_typeCOff3DPoint";   // End point of command
      circleMode : DInt;   // 0: auxPoint defines point on circle line; 1: auxPoint defines circle center; 2: radius and endPoint define circle segment
      circleCenterPoint : "LKinCtrl_typeCOff3DPoint";   // Center point of circle
      circleIntermediatePoint : "LKinCtrl_typeCOff3DPoint";   // Intermediate point of circle
      circleRadius : LReal;   // Radius of circle
      circleAngle : LReal;   // Angle of circle
      pathChoice : DInt;   // circMode(0): not relevant; circMode(1): 0: pos direction; 1: neg direction; circMode(2): 0: short pos segment; 1: short neg segment; 2: long pos segment; 3: long neg segment
      circlePlane : DInt;   // circMode(0): not relevant; circMode(1+2): 0: XZ; 1: YZ; 2: XY
      transitionParameter1 : LReal;   // Transition parameter
      bufferMode : DInt;   // 1: standstill between commands, 2: blending with lower speed; 5: blending with higher speed
   END_STRUCT;
END_TYPE

TYPE "LKinCtrl_typeCOffInCurrentPos"
   STRUCT
      positionAbsolute : "LKinCtrl_typeCartesianPosition";   // Source data - current absolute position
      positionAbsoluteRadComp : "LKinCtrl_typeCartesianPosition";   // Source data - current absolute position radius compensated
   END_STRUCT;
END_TYPE

TYPE "LKinCtrl_typeCOffCmdOutInternal"
   STRUCT
      cmdType : Int := -1;   // 1: MoveLinAbs; 2: MoveLinRel; 3: MoveCircAbs; 4: MoveCircRel; 5: MoveDirectAbs; 6: MoveDirectRel; 10: TrackConveyorBelt; 100: WaitTime; 40/41/42: ContourOffset; 0: FlagOnlyCmd; -1: End of List
      endPoint : "LKinCtrl_typeCOff3DPoint";   // end point of command
      circleMode : DInt;   // 0: auxPoint defines point on circle line; 1: auxPoint defines circle center; 2: radius and endPoint define circle segment
      circleCenterPoint : "LKinCtrl_typeCOff3DPoint";   // center point of circle
      circleIntermediatePoint : "LKinCtrl_typeCOff3DPoint";   // intermediate point of circle
      transitionParameter1 : LReal;   // transition parameter
      endPointOrthShifted : "LKinCtrl_typeCOff3DPoint";   // orthogonal shifted end point of command
      endPointOrthTangShifted : "LKinCtrl_typeCOff3DPoint";   // orthogonal and tangential shifted end point of command
      startPointOrthShifted : "LKinCtrl_typeCOff3DPoint";   // orthogonal shifted end point of command
      startPointOrthTangShifted : "LKinCtrl_typeCOff3DPoint";   // orthogonal and tangential shifted end point of command
      circleRadius : LReal;   // circle radius
      circleAngle : LReal;   // circle angle
      orthogonalUnitVecEnd : "LKinCtrl_typeCOff3DPoint";   // orthogonal unit vector end
      tangentialUnitVecEnd : "LKinCtrl_typeCOff3DPoint";   // tangential unit vector end
      orthogonalShiftEnd : "LKinCtrl_typeCOff3DPoint";   // orthogonal shift end
      tangentiaShiftEnd : "LKinCtrl_typeCOff3DPoint";   // tangential shift end
      orthogonalUnitVecStart : "LKinCtrl_typeCOff3DPoint";   // orthogonal unit vector start
      tangentialUnitVecStart : "LKinCtrl_typeCOff3DPoint";   // tangential unit vector start
      orthogonalShiftStart : "LKinCtrl_typeCOff3DPoint";   // orthogonal shift start
      tangentiaShiftStart : "LKinCtrl_typeCOff3DPoint";   // tangential shift start
      orthogonalUnitVecIntermediate : "LKinCtrl_typeCOff3DPoint";   // orthogonal unit vector intermediate
      tangentialUnitVecIntermediate : "LKinCtrl_typeCOff3DPoint";   // tangential unit vector intermediate
      orthogonalShiftIntermediate : "LKinCtrl_typeCOff3DPoint";   // orthogonal shift intermediate
   END_STRUCT;
END_TYPE

TYPE "LKinCtrl_typeCOffPathDataOut"
   STRUCT
      nextCommand : "LKinCtrl_typePathDataElement";   // Target data - next command
      intermediateCommand : "LKinCtrl_typePathDataElement";   // Target data - intermediate (additional) command
      nextButOneCommand : "LKinCtrl_typeCOffOutNextButOneCmd";   // Target data - next but one command
      nextPositionAbsolute : "LKinCtrl_typeCartesianPosition";   // Source data - next absolute position
      nextPositionAbsoluteRadComp : "LKinCtrl_typeCartesianPosition";   // Source data - next absolute position (radius compensated)
   END_STRUCT;
END_TYPE

// folder: LKinLang_Types

TYPE "LKinLang_typeFileHandlerDiagnostics"
TITLE = typeDiagnosticsFBTemplate
   STRUCT
      status : Word;   // Status of the FB or error identification when error occurred
      subfunctionStatus : Word;   // Status or return value of called FBs, FCs and system blocks
      stateNumber : DInt;   // State in the state machine of the FB when the error occurred
   END_STRUCT;
END_TYPE

TYPE "LKinLang_typeUserDefinedDefaults"
   STRUCT
      velocityLin : LReal := -1.0;   // default velocity for Lin command
   END_STRUCT;
END_TYPE

TYPE "LKinLang_typeVarRef"
   STRUCT
      "name" : String;   // Name of variable
      "type" : Int;   // Type of variable (Local / Interface)
      index : Int;   // Index of variable
      scope : Int;   // Scope of variable (Global / Main / Subprogram)
   END_STRUCT;
END_TYPE

TYPE "LKinLang_typeFileInfo"
   STRUCT
      fileName : String;   // Name of file
      fileState : DInt := 100;   // Actual file status
   END_STRUCT;
END_TYPE

TYPE "LKinLang_typeInterfaceVariables"
   STRUCT
      Boolean : Array[1.."LKINLANG_NUMBER_OF_INTERFACE_BOOL"] of Bool;   // Array of Boolean
      DInts : Array[1.."LKINLANG_NUMBER_OF_INTERFACE_DINT"] of DInt;   // Array of DInt
      LReals : Array[1.."LKINLANG_NUMBER_OF_INTERFACE_LREAL"] of LReal;   // Array of LReal
   END_STRUCT;
END_TYPE

TYPE "LKinLang_typeLabel"
   STRUCT
      lineNumber : UDInt;   // Line number of label
      labelName : String;   // Name of label
      hierarchicLevel : Int;   // Hierarchic level of label
   END_STRUCT;
END_TYPE

TYPE "LKinLang_typeLabelList"
   STRUCT
      numberOfLabels : Int;   // Counter of found labels
      labels : Array[1.."LKINLANG_NUMBER_OF_LABELS"] of "LKinLang_typeLabel";   // Array of labels
   END_STRUCT;
END_TYPE

TYPE "LKinLang_typeVarRefList"
   STRUCT
      numberOfReferences : Int;   // Number of variable references
      references : Array[1.."LKINLANG_NUMBER_OF_VAR_REFS"] of "LKinLang_typeVarRef";   // Array of references
   END_STRUCT;
END_TYPE

TYPE "LKinLang_typeLocalVariables"
   STRUCT
      boolCounter : Int;   // Number of boolean variables
      dintCounter : Int;   // Number of integer variables
      lrealCounter : Int;   // Number of real variables
      boolean : Array[1.."LKINLANG_NUMBER_OF_LOCAL_BOOL"] of Bool;   // Array of loca boolean
      dints : Array[1.."LKINLANG_NUMBER_OF_LOCAL_DINT"] of DInt;   // Array of local integer
      lreals : Array[1.."LKINLANG_NUMBER_OF_LOCAL_LREAL"] of LReal;   // Array of local real
   END_STRUCT;
END_TYPE

TYPE "LKinLang_typeLocalVarDefinition"
   STRUCT
      tokenizedString : "LKinLang_typeLineTokens";   // Tokenized string
      nameTokenNumber : USInt;   // Index of the "_name_" token
      typeTokenNumber : USInt;   // Index of the "_type_" token
   END_STRUCT;
END_TYPE

TYPE "LKinLang_typeLineBufferPointer"
VERSION : 0.1
   STRUCT
      addPointer : DInt := 0;   // pointer to add new comds to PathData after cmd has been executed by MovePath
      retrievePointer : DInt := 0;   // pointer to show which cmd is the next to be retrieved by MovePath
      addPointerRestarted : Bool;   // addPointer restarted after overflow
      ignoreAddPointer : Bool := true;   // addPointer not taken into account for buffering, unless set by previous data source
      bufferLocked : Bool;   // buffer locked to wait for previous data source - read data locked
      endOfFile : Bool;   // end of file reached
      restart : Bool;   // restart reading file; set by parser
      requestedLine : UDInt;   // Parser can request line number here for jumps
   END_STRUCT;
END_TYPE
